REGION Network 11: Motor Conveyor Labeller
   RUNG wire#powerrail
      Contact( "Flag Motor" )
      Coil( "Motor" )
   END_RUNG
   // the same network as SCL:
   "Motor" := "Flag Motor";
END_REGION

REGION Network 12: Start Markem Input
   RUNG wire#powerrail
      Contact( "Flag Imaje Start" )
      Coil( "Imaje Output Start" )
   END_RUNG
   // the same network as SCL:
   "Imaje Output Start" := "Flag Imaje Start";
END_REGION

REGION Network 13: Pause Markem Input
   RUNG wire#powerrail
      Contact( "Flag Imaje Pause" )
      Coil( "Imaje Output Pause" )
   END_RUNG
   // the same network as SCL:
   "Imaje Output Pause" := "Flag Imaje Pause";
END_REGION

REGION Network 14: Trigger Markem Stamp
   RUNG wire#powerrail
      Contact( "Flag Imaje Trigger" )
      Coil( "Imaje Output Trigger" )
   END_RUNG
   // the same network as SCL:
   "Imaje Output Trigger" := "Flag Imaje Trigger";
END_REGION

REGION Network 15: Mesin Sebelumnya
   RUNG wire#powerrail
      Contact( "Machine Running" )
      Coil( "Trigger Mesin Sebelumnya" )
   END_RUNG
   // the same network as SCL:
   "Trigger Mesin Sebelumnya" := "Machine Running";
END_REGION

REGION Network 16: Error Output
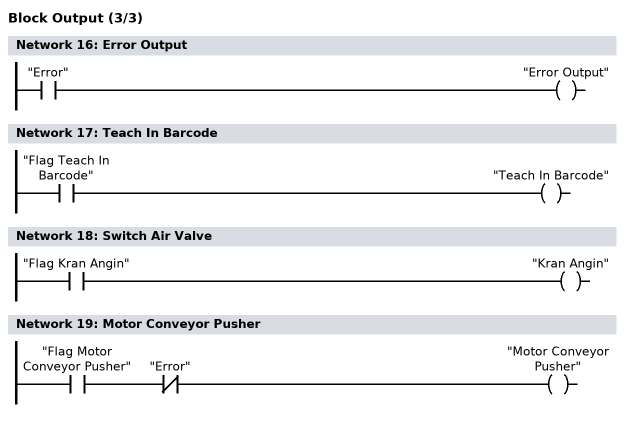
   RUNG wire#powerrail
      Contact( "Error" )
      Coil( "Error Output" )
   END_RUNG
   // the same network as SCL:
   "Error Output" := "Error";
END_REGION

REGION Network 17: Teach In Barcode
   RUNG wire#powerrail
      Contact( "Flag Teach In Barcode" )
      Coil( "Teach In Barcode" )
   END_RUNG
   // the same network as SCL:
   "Teach In Barcode" := "Flag Teach In Barcode";
END_REGION

REGION Network 18: Switch Air Valve
   RUNG wire#powerrail
      Contact( "Flag Kran Angin" )
      Coil( "Kran Angin" )
   END_RUNG
   // the same network as SCL:
   "Kran Angin" := "Flag Kran Angin";
END_REGION

REGION Network 19: Motor Conveyor Pusher
   RUNG wire#powerrail
      Contact( "Flag Motor Conveyor Pusher" )
      I_Contact( "Error" )
      Coil( "Motor Conveyor Pusher" )
   END_RUNG
   // the same network as SCL:
   "Motor Conveyor Pusher" := "Flag Motor Conveyor Pusher" AND NOT "Error";
END_REGION

REGION Network 20: Motor Heating Roll
END_REGION
END_FUNCTION_BLOCK

FUNCTION_BLOCK "S Block Current Shift"   // FB4, LAD
{ S7_Optimized_Access := 'TRUE' }
VERSION : 0.1
   VAR_TEMP   // added for the SCL form of the ladder/FBD networks
      _w1 : Bool;
      _w2 : Bool;
   END_VAR
BEGIN

REGION Network 1: Input Sloft ........................................................................page 1
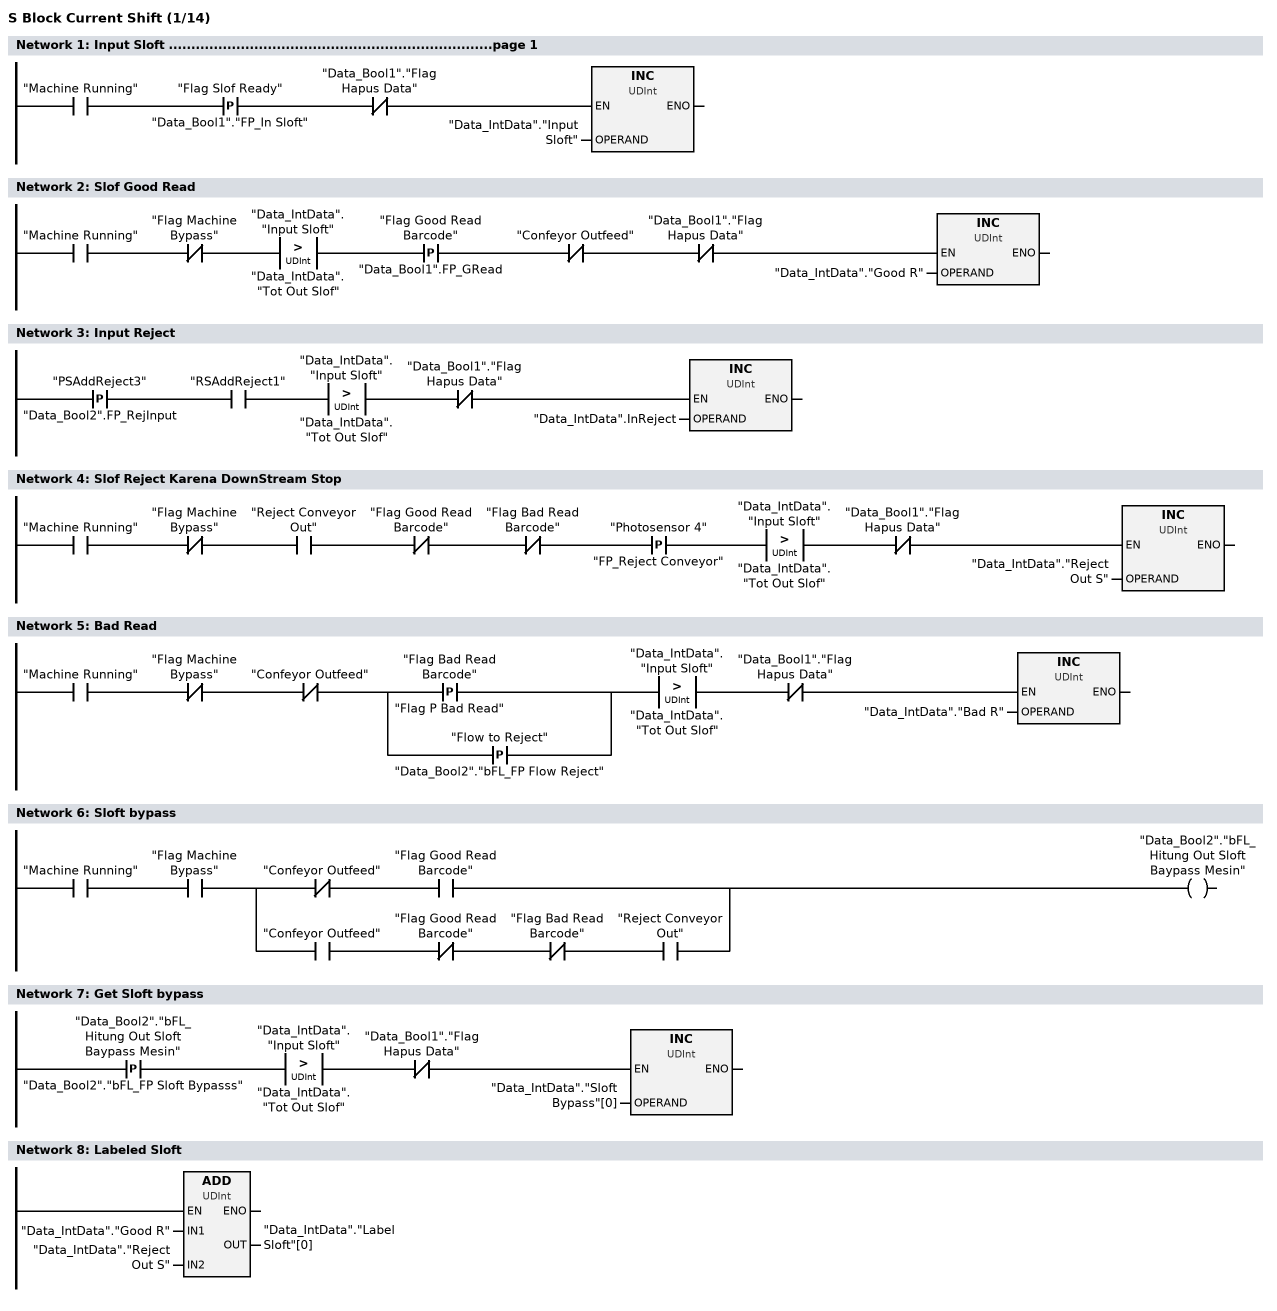
   RUNG wire#powerrail
      Contact( "Machine Running" )
      P_Contact(operand := "Flag Slof Ready", bit := "Data_Bool1"."FP_In Sloft")
      I_Contact( "Data_Bool1"."Flag Hapus Data" )
      { S7_Templates := "DestType := UDInt"; S7_GenerateENO := "TRUE" } Inc( "Data_IntData"."Input Sloft" )
   END_RUNG
   // the same network as SCL:
   #_w1 := "Machine Running" AND "Flag Slof Ready" AND NOT "Data_Bool1"."FP_In Sloft";   // rising edge of "Flag Slof Ready"
   "Data_Bool1"."FP_In Sloft" := "Flag Slof Ready";
   IF #_w1 AND NOT "Data_Bool1"."Flag Hapus Data" THEN
       "Data_IntData"."Input Sloft" := "Data_IntData"."Input Sloft" + 1;
   END_IF;
END_REGION

REGION Network 2: Slof Good Read
   RUNG wire#powerrail
      Contact( "Machine Running" )
      I_Contact( "Flag Machine Bypass" )
      { S7_Templates := "SrcType := UDInt" } GT_Contact(in1 := "Data_IntData"."Input Sloft", in2 := "Data_IntData"."Tot Out Slof")
      P_Contact(operand := "Flag Good Read Barcode", bit := "Data_Bool1".FP_GRead)
      I_Contact( "Confeyor Outfeed" )
      I_Contact( "Data_Bool1"."Flag Hapus Data" )
      { S7_Templates := "DestType := UDInt"; S7_GenerateENO := "TRUE" } Inc( "Data_IntData"."Good R" )
   END_RUNG
   // the same network as SCL:
   #_w1 := "Machine Running" AND NOT "Flag Machine Bypass" AND ("Data_IntData"."Input Sloft" > "Data_IntData"."Tot Out Slof") AND "Flag Good Read Barcode" AND NOT "Data_Bool1".FP_GRead;   // rising edge of "Flag Good Read Barcode"
   "Data_Bool1".FP_GRead := "Flag Good Read Barcode";
   IF #_w1 AND NOT "Confeyor Outfeed" AND NOT "Data_Bool1"."Flag Hapus Data" THEN
       "Data_IntData"."Good R" := "Data_IntData"."Good R" + 1;
   END_IF;
END_REGION

REGION Network 3: Input Reject
   RUNG wire#powerrail
      P_Contact(operand := "PSAddReject3", bit := "Data_Bool2".FP_RejInput)
      Contact( "RSAddReject1" )
      { S7_Templates := "SrcType := UDInt" } GT_Contact(in1 := "Data_IntData"."Input Sloft", in2 := "Data_IntData"."Tot Out Slof")
      I_Contact( "Data_Bool1"."Flag Hapus Data" )
      { S7_Templates := "DestType := UDInt"; S7_GenerateENO := "TRUE" } Inc( "Data_IntData".InReject )
   END_RUNG
   // the same network as SCL:
   #_w1 := "PSAddReject3" AND NOT "Data_Bool2".FP_RejInput;   // rising edge of "PSAddReject3"
   "Data_Bool2".FP_RejInput := "PSAddReject3";
   IF #_w1 AND "RSAddReject1" AND ("Data_IntData"."Input Sloft" > "Data_IntData"."Tot Out Slof") AND NOT "Data_Bool1"."Flag Hapus Data" THEN
       "Data_IntData".InReject := "Data_IntData".InReject + 1;
   END_IF;
END_REGION

REGION Network 4: Slof Reject Karena DownStream Stop
   RUNG wire#powerrail
      Contact( "Machine Running" )
      I_Contact( "Flag Machine Bypass" )
      Contact( "Reject Conveyor Out" )
      I_Contact( "Flag Good Read Barcode" )
      I_Contact( "Flag Bad Read Barcode" )
      P_Contact(operand := "Photosensor 4", bit := "FP_Reject Conveyor")
      { S7_Templates := "SrcType := UDInt" } GT_Contact(in1 := "Data_IntData"."Input Sloft", in2 := "Data_IntData"."Tot Out Slof")
      I_Contact( "Data_Bool1"."Flag Hapus Data" )
      { S7_Templates := "DestType := UDInt"; S7_GenerateENO := "TRUE" } Inc( "Data_IntData"."Reject Out S" )
   END_RUNG
   // the same network as SCL:
   #_w1 := "Machine Running" AND NOT "Flag Machine Bypass" AND "Reject Conveyor Out" AND NOT "Flag Good Read Barcode" AND NOT "Flag Bad Read Barcode" AND "Photosensor 4" AND NOT "FP_Reject Conveyor";   // rising edge of "Photosensor 4"
   "FP_Reject Conveyor" := "Photosensor 4";
   IF #_w1 AND ("Data_IntData"."Input Sloft" > "Data_IntData"."Tot Out Slof") AND NOT "Data_Bool1"."Flag Hapus Data" THEN
       "Data_IntData"."Reject Out S" := "Data_IntData"."Reject Out S" + 1;
   END_IF;
END_REGION

REGION Network 5: Bad Read
   RUNG wire#powerrail
      Contact( "Machine Running" )
      I_Contact( "Flag Machine Bypass" )
      I_Contact( "Confeyor Outfeed" )
      wire#w1
      P_Contact(operand := "Flag Bad Read Barcode", bit := "Flag P Bad Read")
      wire#w2
      { S7_Templates := "SrcType := UDInt" } GT_Contact(in1 := "Data_IntData"."Input Sloft", in2 := "Data_IntData"."Tot Out Slof")
      I_Contact( "Data_Bool1"."Flag Hapus Data" )
      { S7_Templates := "DestType := UDInt"; S7_GenerateENO := "TRUE" } Inc( "Data_IntData"."Bad R" )
   END_RUNG
   RUNG wire#w1
      P_Contact(operand := "Flow to Reject", bit := "Data_Bool2"."bFL_FP Flow Reject")
   END_RUNG wire#w2
   // the same network as SCL:
   #_w1 := "Machine Running" AND NOT "Flag Machine Bypass" AND NOT "Confeyor Outfeed" AND "Flag Bad Read Barcode" AND NOT "Flag P Bad Read";   // rising edge of "Flag Bad Read Barcode"
   "Flag P Bad Read" := "Flag Bad Read Barcode";
   #_w2 := "Machine Running" AND NOT "Flag Machine Bypass" AND NOT "Confeyor Outfeed" AND "Flow to Reject" AND NOT "Data_Bool2"."bFL_FP Flow Reject";   // rising edge of "Flow to Reject"
   "Data_Bool2"."bFL_FP Flow Reject" := "Flow to Reject";
   IF (#_w1 OR #_w2) AND ("Data_IntData"."Input Sloft" > "Data_IntData"."Tot Out Slof") AND NOT "Data_Bool1"."Flag Hapus Data" THEN
       "Data_IntData"."Bad R" := "Data_IntData"."Bad R" + 1;
   END_IF;
END_REGION

REGION Network 6: Sloft bypass
   RUNG wire#powerrail
      Contact( "Machine Running" )
      Contact( "Flag Machine Bypass" )
      wire#w1
      I_Contact( "Confeyor Outfeed" )
      Contact( "Flag Good Read Barcode" )
      wire#w2
      Coil( "Data_Bool2"."bFL_Hitung Out Sloft Baypass Mesin" )
   END_RUNG
   RUNG wire#w1
      Contact( "Confeyor Outfeed" )
      I_Contact( "Flag Good Read Barcode" )
      I_Contact( "Flag Bad Read Barcode" )
      Contact( "Reject Conveyor Out" )
   END_RUNG wire#w2
   // the same network as SCL:
   "Data_Bool2"."bFL_Hitung Out Sloft Baypass Mesin" := "Machine Running" AND "Flag Machine Bypass" AND ((NOT "Confeyor Outfeed" AND "Flag Good Read Barcode") OR ("Confeyor Outfeed" AND NOT "Flag Good Read Barcode" AND NOT "Flag Bad Read Barcode" AND "Reject Conveyor Out"));
END_REGION

REGION Network 7: Get Sloft bypass
   RUNG wire#powerrail
      P_Contact(operand := "Data_Bool2"."bFL_Hitung Out Sloft Baypass Mesin", bit := "Data_Bool2"."bFL_FP Sloft Bypasss")
      { S7_Templates := "SrcType := UDInt" } GT_Contact(in1 := "Data_IntData"."Input Sloft", in2 := "Data_IntData"."Tot Out Slof")
      I_Contact( "Data_Bool1"."Flag Hapus Data" )
      { S7_Templates := "DestType := UDInt"; S7_GenerateENO := "TRUE" } Inc( "Data_IntData"."Sloft Bypass"[0] )
   END_RUNG
   // the same network as SCL:
   #_w1 := "Data_Bool2"."bFL_Hitung Out Sloft Baypass Mesin" AND NOT "Data_Bool2"."bFL_FP Sloft Bypasss";   // rising edge of "Data_Bool2"."bFL_Hitung Out Sloft Baypass Mesin"
   "Data_Bool2"."bFL_FP Sloft Bypasss" := "Data_Bool2"."bFL_Hitung Out Sloft Baypass Mesin";
   IF #_w1 AND ("Data_IntData"."Input Sloft" > "Data_IntData"."Tot Out Slof") AND NOT "Data_Bool1"."Flag Hapus Data" THEN
       "Data_IntData"."Sloft Bypass"[0] := "Data_IntData"."Sloft Bypass"[0] + 1;
   END_IF;
END_REGION

REGION Network 8: Labeled Sloft
   RUNG wire#powerrail
      { S7_Templates := "SrcType := UDInt"; S7_GenerateENO := "TRUE" } Add(in1 := "Data_IntData"."Good R", in2 := "Data_IntData"."Reject Out S", out => "Data_IntData"."Label Sloft"[0])
   END_RUNG
   // the same network as SCL:
   "Data_IntData"."Label Sloft"[0] := "Data_IntData"."Good R" + "Data_IntData"."Reject Out S";
END_REGION

REGION Network 9: Unlabeled Sloft
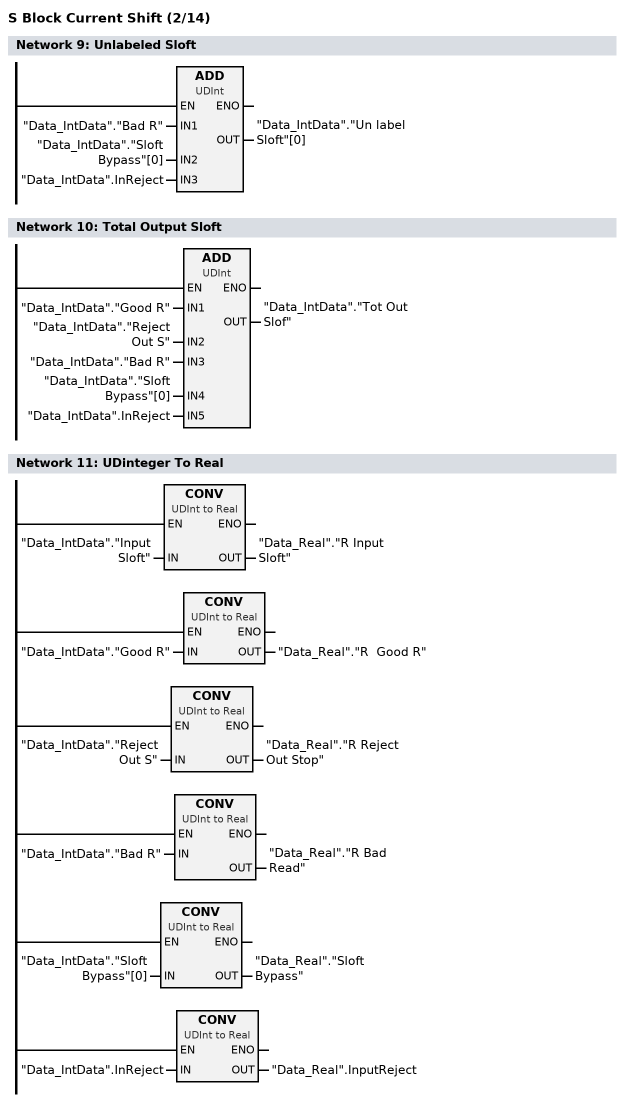
   RUNG wire#powerrail
      { S7_Templates := "SrcType := UDInt"; S7_GenerateENO := "TRUE" } Add(in1 := "Data_IntData"."Bad R", in2 := "Data_IntData"."Sloft Bypass"[0], in3 := "Data_IntData".InReject, out => "Data_IntData"."Un label Sloft"[0])
   END_RUNG
   // the same network as SCL:
   "Data_IntData"."Un label Sloft"[0] := "Data_IntData"."Bad R" + "Data_IntData"."Sloft Bypass"[0] + "Data_IntData".InReject;
END_REGION

REGION Network 10: Total Output Sloft
   RUNG wire#powerrail
      { S7_Templates := "SrcType := UDInt"; S7_GenerateENO := "TRUE" } Add(in1 := "Data_IntData"."Good R", in2 := "Data_IntData"."Reject Out S", in3 := "Data_IntData"."Bad R", in4 := "Data_IntData"."Sloft Bypass"[0], in5 := "Data_IntData".InReject, out => "Data_IntData"."Tot Out Slof")
   END_RUNG
   // the same network as SCL:
   "Data_IntData"."Tot Out Slof" := "Data_IntData"."Good R" + "Data_IntData"."Reject Out S" + "Data_IntData"."Bad R" + "Data_IntData"."Sloft Bypass"[0] + "Data_IntData".InReject;
END_REGION

REGION Network 11: UDinteger To Real
   RUNG wire#powerrail
      { S7_Templates := "[SrcType := UDInt, DestType := Real]"; S7_GenerateENO := "TRUE" } Convert(in := "Data_IntData"."Input Sloft", out => "Data_Real"."R Input Sloft")
   END_RUNG
   RUNG wire#powerrail
      { S7_Templates := "[SrcType := UDInt, DestType := Real]"; S7_GenerateENO := "TRUE" } Convert(in := "Data_IntData"."Good R", out => "Data_Real"."R  Good R")
   END_RUNG
   RUNG wire#powerrail
      { S7_Templates := "[SrcType := UDInt, DestType := Real]"; S7_GenerateENO := "TRUE" } Convert(in := "Data_IntData"."Reject Out S", out => "Data_Real"."R Reject Out Stop")
   END_RUNG
   RUNG wire#powerrail
      { S7_Templates := "[SrcType := UDInt, DestType := Real]"; S7_GenerateENO := "TRUE" } Convert(in := "Data_IntData"."Bad R", out => "Data_Real"."R Bad Read")
   END_RUNG
   RUNG wire#powerrail
      { S7_Templates := "[SrcType := UDInt, DestType := Real]"; S7_GenerateENO := "TRUE" } Convert(in := "Data_IntData"."Sloft Bypass"[0], out => "Data_Real"."Sloft Bypass")
   END_RUNG
   RUNG wire#powerrail
      { S7_Templates := "[SrcType := UDInt, DestType := Real]"; S7_GenerateENO := "TRUE" } Convert(in := "Data_IntData".InReject, out => "Data_Real".InputReject)
   END_RUNG
   // the same network as SCL:
   "Data_Real"."R Input Sloft" := UDINT_TO_REAL("Data_IntData"."Input Sloft");
   "Data_Real"."R  Good R" := UDINT_TO_REAL("Data_IntData"."Good R");
   "Data_Real"."R Reject Out Stop" := UDINT_TO_REAL("Data_IntData"."Reject Out S");
   "Data_Real"."R Bad Read" := UDINT_TO_REAL("Data_IntData"."Bad R");
   "Data_Real"."Sloft Bypass" := UDINT_TO_REAL("Data_IntData"."Sloft Bypass"[0]);
   "Data_Real".InputReject := UDINT_TO_REAL("Data_IntData".InReject);
END_REGION

REGION Network 12: % Sloft terhadap Input Sloft
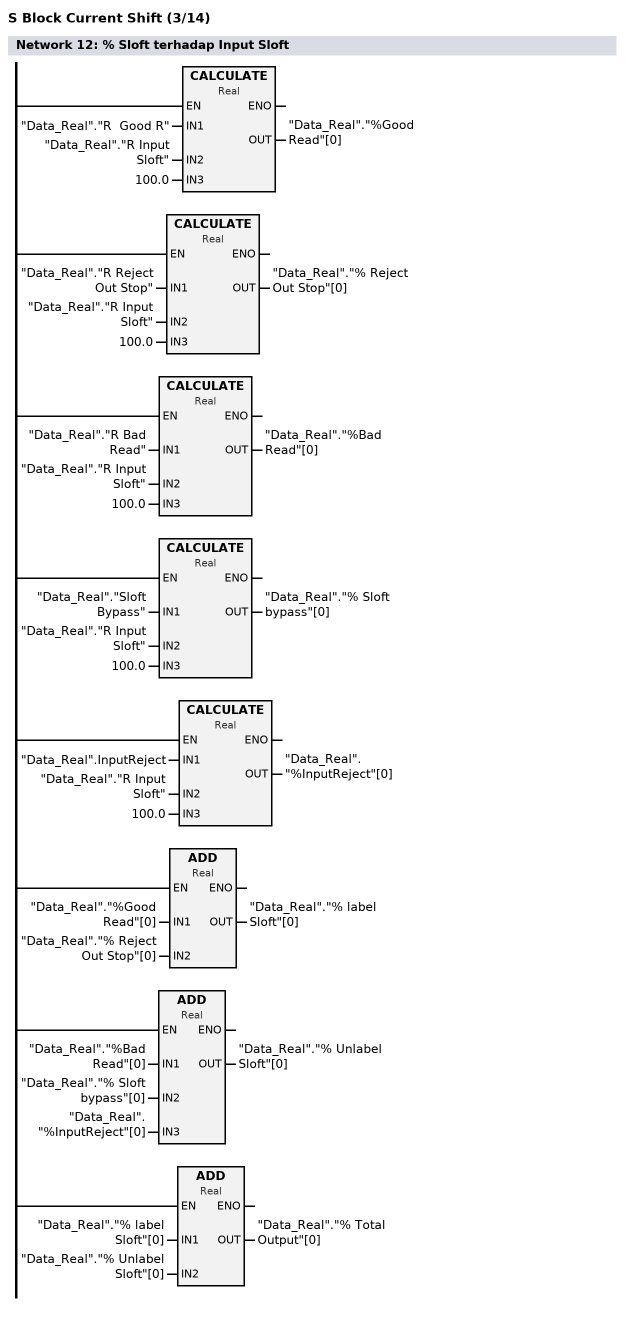
   RUNG wire#powerrail
      { S7_Templates := "SrcType := Real"; S7_GenerateENO := "TRUE"; S7_Expression := "(IN1/IN2)*IN3" } Calculate(in1 := "Data_Real"."R  Good R", in2 := "Data_Real"."R Input Sloft", in3 := 100.0, out => "Data_Real"."%Good Read"[0])
   END_RUNG
   RUNG wire#powerrail
      { S7_Templates := "SrcType := Real"; S7_GenerateENO := "TRUE"; S7_Expression := "(IN1/IN2)*IN3" } Calculate(in1 := "Data_Real"."R Reject Out Stop", in2 := "Data_Real"."R Input Sloft", in3 := 100.0, out => "Data_Real"."% Reject Out Stop"[0])
   END_RUNG
   RUNG wire#powerrail
      { S7_Templates := "SrcType := Real"; S7_GenerateENO := "TRUE"; S7_Expression := "(IN1/IN2)*IN3" } Calculate(in1 := "Data_Real"."R Bad Read", in2 := "Data_Real"."R Input Sloft", in3 := 100.0, out => "Data_Real"."%Bad Read"[0])
   END_RUNG
   RUNG wire#powerrail
      { S7_Templates := "SrcType := Real"; S7_GenerateENO := "TRUE"; S7_Expression := "(IN1/IN2)*IN3" } Calculate(in1 := "Data_Real"."Sloft Bypass", in2 := "Data_Real"."R Input Sloft", in3 := 100.0, out => "Data_Real"."% Sloft bypass"[0])
   END_RUNG
   RUNG wire#powerrail
      { S7_Templates := "SrcType := Real"; S7_GenerateENO := "TRUE"; S7_Expression := "(IN1/IN2)*IN3" } Calculate(in1 := "Data_Real".InputReject, in2 := "Data_Real"."R Input Sloft", in3 := 100.0, out => "Data_Real"."%InputReject"[0])
   END_RUNG
   RUNG wire#powerrail
      { S7_Templates := "SrcType := Real"; S7_GenerateENO := "TRUE" } Add(in1 := "Data_Real"."%Good Read"[0], in2 := "Data_Real"."% Reject Out Stop"[0], out => "Data_Real"."% label Sloft"[0])
   END_RUNG
   RUNG wire#powerrail
      { S7_Templates := "SrcType := Real"; S7_GenerateENO := "TRUE" } Add(in1 := "Data_Real"."%Bad Read"[0], in2 := "Data_Real"."% Sloft bypass"[0], in3 := "Data_Real"."%InputReject"[0], out => "Data_Real"."% Unlabel Sloft"[0])
   END_RUNG
   RUNG wire#powerrail
      { S7_Templates := "SrcType := Real"; S7_GenerateENO := "TRUE" } Add(in1 := "Data_Real"."% label Sloft"[0], in2 := "Data_Real"."% Unlabel Sloft"[0], out => "Data_Real"."% Total Output"[0])
   END_RUNG
   // the same network as SCL:
   "Data_Real"."%Good Read"[0] := ("Data_Real"."R  Good R"/"Data_Real"."R Input Sloft")*100.0;
   "Data_Real"."% Reject Out Stop"[0] := ("Data_Real"."R Reject Out Stop"/"Data_Real"."R Input Sloft")*100.0;
   "Data_Real"."%Bad Read"[0] := ("Data_Real"."R Bad Read"/"Data_Real"."R Input Sloft")*100.0;
   "Data_Real"."% Sloft bypass"[0] := ("Data_Real"."Sloft Bypass"/"Data_Real"."R Input Sloft")*100.0;
   "Data_Real"."%InputReject"[0] := ("Data_Real".InputReject/"Data_Real"."R Input Sloft")*100.0;
   "Data_Real"."% label Sloft"[0] := "Data_Real"."%Good Read"[0] + "Data_Real"."% Reject Out Stop"[0];
   "Data_Real"."% Unlabel Sloft"[0] := "Data_Real"."%Bad Read"[0] + "Data_Real"."% Sloft bypass"[0] + "Data_Real"."%InputReject"[0];
   "Data_Real"."% Total Output"[0] := "Data_Real"."% label Sloft"[0] + "Data_Real"."% Unlabel Sloft"[0];
END_REGION

REGION Network 13: ----------- Get Image Output Trigger
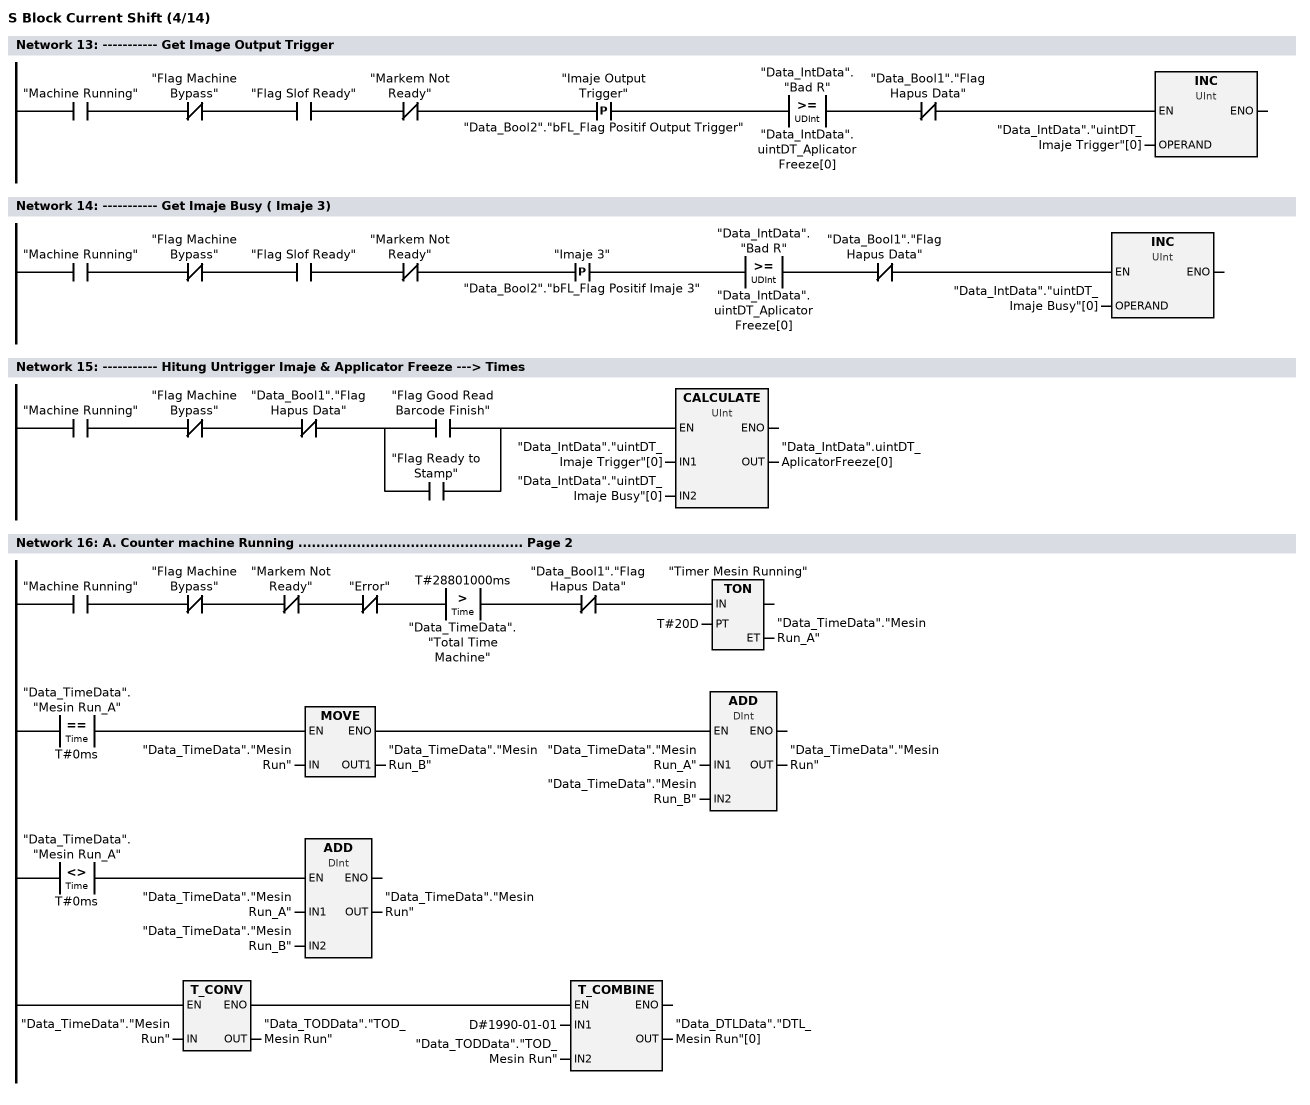
   RUNG wire#powerrail
      Contact( "Machine Running" )
      I_Contact( "Flag Machine Bypass" )
      Contact( "Flag Slof Ready" )
      I_Contact( "Markem Not Ready" )
      P_Contact(operand := "Imaje Output Trigger", bit := "Data_Bool2"."bFL_Flag Positif Output Trigger")
      { S7_Templates := "SrcType := UDInt" } GE_Contact(in1 := "Data_IntData"."Bad R", in2 := "Data_IntData".uintDT_AplicatorFreeze[0])
      I_Contact( "Data_Bool1"."Flag Hapus Data" )
      { S7_Templates := "DestType := UInt"; S7_GenerateENO := "TRUE" } Inc( "Data_IntData"."uintDT_Imaje Trigger"[0] )
   END_RUNG
   // the same network as SCL:
   #_w1 := "Machine Running" AND NOT "Flag Machine Bypass" AND "Flag Slof Ready" AND NOT "Markem Not Ready" AND "Imaje Output Trigger" AND NOT "Data_Bool2"."bFL_Flag Positif Output Trigger";   // rising edge of "Imaje Output Trigger"
   "Data_Bool2"."bFL_Flag Positif Output Trigger" := "Imaje Output Trigger";
   IF #_w1 AND ("Data_IntData"."Bad R" >= "Data_IntData".uintDT_AplicatorFreeze[0]) AND NOT "Data_Bool1"."Flag Hapus Data" THEN
       "Data_IntData"."uintDT_Imaje Trigger"[0] := "Data_IntData"."uintDT_Imaje Trigger"[0] + 1;
   END_IF;
END_REGION

REGION Network 14: ----------- Get Imaje Busy ( Imaje 3)
   RUNG wire#powerrail
      Contact( "Machine Running" )
      I_Contact( "Flag Machine Bypass" )
      Contact( "Flag Slof Ready" )
      I_Contact( "Markem Not Ready" )
      P_Contact(operand := "Imaje 3", bit := "Data_Bool2"."bFL_Flag Positif Imaje 3")
      { S7_Templates := "SrcType := UDInt" } GE_Contact(in1 := "Data_IntData"."Bad R", in2 := "Data_IntData".uintDT_AplicatorFreeze[0])
      I_Contact( "Data_Bool1"."Flag Hapus Data" )
      { S7_Templates := "DestType := UInt"; S7_GenerateENO := "TRUE" } Inc( "Data_IntData"."uintDT_Imaje Busy"[0] )
   END_RUNG
   // the same network as SCL:
   #_w1 := "Machine Running" AND NOT "Flag Machine Bypass" AND "Flag Slof Ready" AND NOT "Markem Not Ready" AND "Imaje 3" AND NOT "Data_Bool2"."bFL_Flag Positif Imaje 3";   // rising edge of "Imaje 3"
   "Data_Bool2"."bFL_Flag Positif Imaje 3" := "Imaje 3";
   IF #_w1 AND ("Data_IntData"."Bad R" >= "Data_IntData".uintDT_AplicatorFreeze[0]) AND NOT "Data_Bool1"."Flag Hapus Data" THEN
       "Data_IntData"."uintDT_Imaje Busy"[0] := "Data_IntData"."uintDT_Imaje Busy"[0] + 1;
   END_IF;
END_REGION

REGION Network 15: ----------- Hitung Untrigger Imaje & Applicator Freeze ---> Times
   RUNG wire#powerrail
      Contact( "Machine Running" )
      I_Contact( "Flag Machine Bypass" )
      I_Contact( "Data_Bool1"."Flag Hapus Data" )
      wire#w1
      Contact( "Flag Good Read Barcode Finish" )
      wire#w2
      { S7_Templates := "SrcType := UInt"; S7_GenerateENO := "TRUE"; S7_Expression := "IN1- IN2" } Calculate(in1 := "Data_IntData"."uintDT_Imaje Trigger"[0], in2 := "Data_IntData"."uintDT_Imaje Busy"[0], out => "Data_IntData".uintDT_AplicatorFreeze[0])
   END_RUNG
   RUNG wire#w1
      Contact( "Flag Ready to Stamp" )
   END_RUNG wire#w2
   // the same network as SCL:
   IF "Machine Running" AND NOT "Flag Machine Bypass" AND NOT "Data_Bool1"."Flag Hapus Data" AND ("Flag Good Read Barcode Finish" OR "Flag Ready to Stamp") THEN
       "Data_IntData".uintDT_AplicatorFreeze[0] := "Data_IntData"."uintDT_Imaje Trigger"[0]- "Data_IntData"."uintDT_Imaje Busy"[0];
   END_IF;
END_REGION

REGION Network 16: A. Counter machine Running .................................................. Page 2
   // ENO of a box is taken as its EN; it also drops when the box reports an error
   "Timer Mesin Running".TON(IN := "Machine Running" AND NOT "Flag Machine Bypass" AND NOT "Markem Not Ready" AND NOT "Error" AND (T#28801000ms > "Data_TimeData"."Total Time Machine") AND NOT "Data_Bool1"."Flag Hapus Data",
                           PT := T#20D,
                           ET => "Data_TimeData"."Mesin Run_A");
   IF "Data_TimeData"."Mesin Run_A" = T#0ms THEN
       "Data_TimeData"."Mesin Run_B" := "Data_TimeData"."Mesin Run";
       "Data_TimeData"."Mesin Run" := "Data_TimeData"."Mesin Run_A" + "Data_TimeData"."Mesin Run_B";
   END_IF;
   IF "Data_TimeData"."Mesin Run_A" <> T#0ms THEN
       "Data_TimeData"."Mesin Run" := "Data_TimeData"."Mesin Run_A" + "Data_TimeData"."Mesin Run_B";
   END_IF;
   "Data_TODData"."TOD_Mesin Run" := T_CONV(IN := "Data_TimeData"."Mesin Run");
   "Data_DTLData"."DTL_Mesin Run"[0] := T_COMBINE(IN1 := D#1990-01-01, IN2 := "Data_TODData"."TOD_Mesin Run");
END_REGION

REGION Network 17: B. Counter machine Running Baypass Stamp
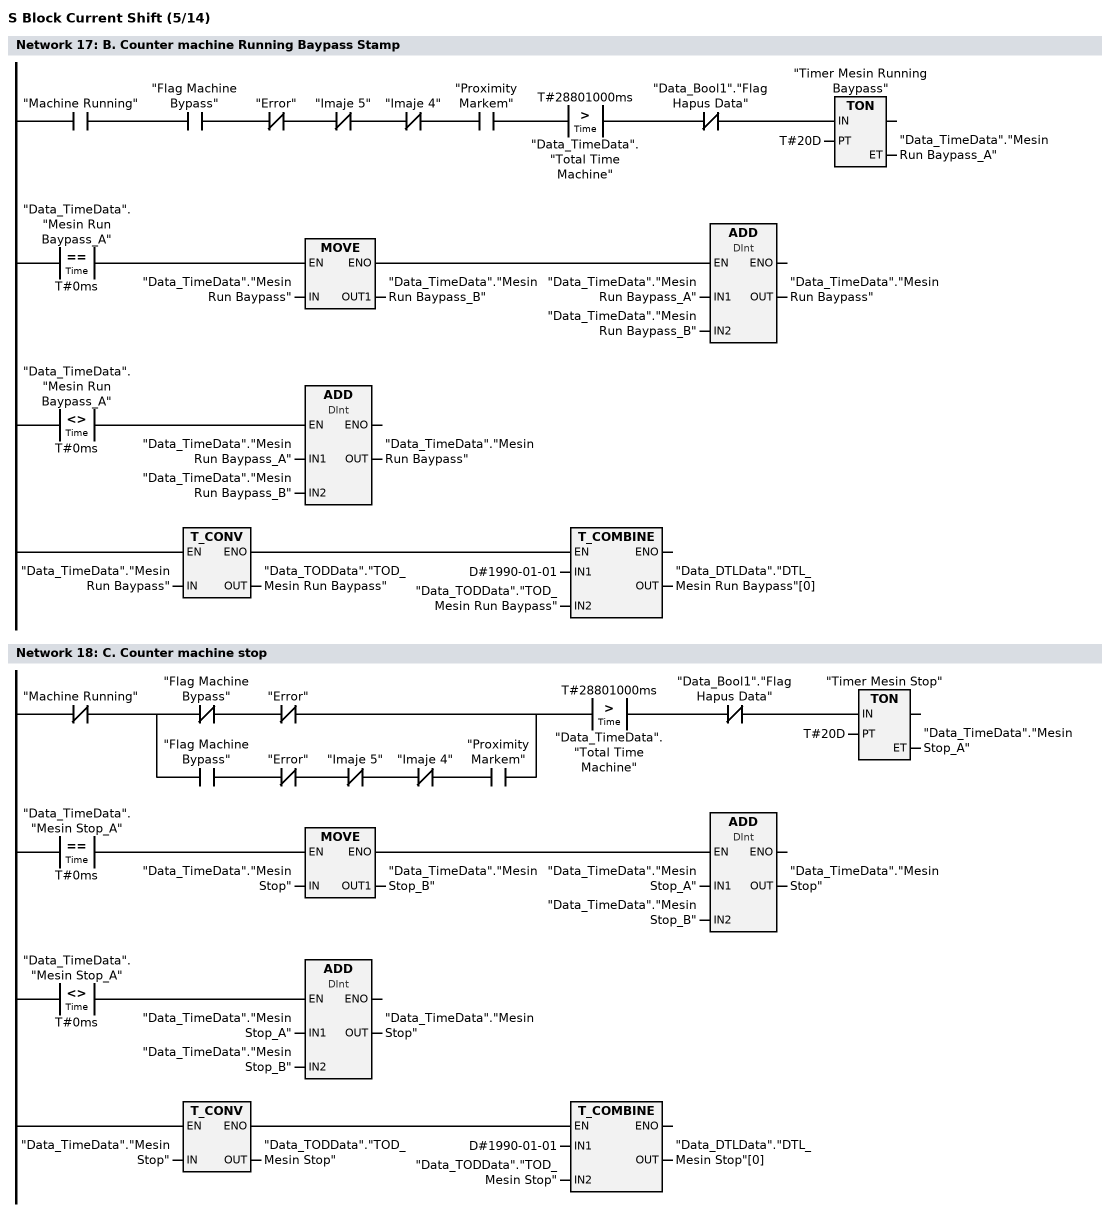
   // ENO of a box is taken as its EN; it also drops when the box reports an error
   "Timer Mesin Running Baypass".TON(IN := "Machine Running" AND "Flag Machine Bypass" AND NOT "Error" AND NOT "Imaje 5" AND NOT "Imaje 4" AND "Proximity Markem" AND (T#28801000ms > "Data_TimeData"."Total Time Machine") AND NOT "Data_Bool1"."Flag Hapus Data",
                           PT := T#20D,
                           ET => "Data_TimeData"."Mesin Run Baypass_A");
   IF "Data_TimeData"."Mesin Run Baypass_A" = T#0ms THEN
       "Data_TimeData"."Mesin Run Baypass_B" := "Data_TimeData"."Mesin Run Baypass";
       "Data_TimeData"."Mesin Run Baypass" := "Data_TimeData"."Mesin Run Baypass_A" + "Data_TimeData"."Mesin Run Baypass_B";
   END_IF;
   IF "Data_TimeData"."Mesin Run Baypass_A" <> T#0ms THEN
       "Data_TimeData"."Mesin Run Baypass" := "Data_TimeData"."Mesin Run Baypass_A" + "Data_TimeData"."Mesin Run Baypass_B";
   END_IF;
   "Data_TODData"."TOD_Mesin Run Baypass" := T_CONV(IN := "Data_TimeData"."Mesin Run Baypass");
   "Data_DTLData"."DTL_Mesin Run Baypass"[0] := T_COMBINE(IN1 := D#1990-01-01,
                           IN2 := "Data_TODData"."TOD_Mesin Run Baypass");
END_REGION

REGION Network 18: C. Counter machine stop
   // ENO of a box is taken as its EN; it also drops when the box reports an error
   "Timer Mesin Stop".TON(IN := NOT "Machine Running" AND ((NOT "Flag Machine Bypass" AND NOT "Error") OR ("Flag Machine Bypass" AND NOT "Error" AND NOT "Imaje 5" AND NOT "Imaje 4" AND "Proximity Markem")) AND (T#28801000ms > "Data_TimeData"."Total Time Machine") AND NOT "Data_Bool1"."Flag Hapus Data",
                          PT := T#20D,
                          ET => "Data_TimeData"."Mesin Stop_A");
   IF "Data_TimeData"."Mesin Stop_A" = T#0ms THEN
       "Data_TimeData"."Mesin Stop_B" := "Data_TimeData"."Mesin Stop";
       "Data_TimeData"."Mesin Stop" := "Data_TimeData"."Mesin Stop_A" + "Data_TimeData"."Mesin Stop_B";
   END_IF;
   IF "Data_TimeData"."Mesin Stop_A" <> T#0ms THEN
       "Data_TimeData"."Mesin Stop" := "Data_TimeData"."Mesin Stop_A" + "Data_TimeData"."Mesin Stop_B";
   END_IF;
   "Data_TODData"."TOD_Mesin Stop" := T_CONV(IN := "Data_TimeData"."Mesin Stop");
   "Data_DTLData"."DTL_Mesin Stop"[0] := T_COMBINE(IN1 := D#1990-01-01, IN2 := "Data_TODData"."TOD_Mesin Stop");
END_REGION

REGION Network 19: D. Counter Machine Error
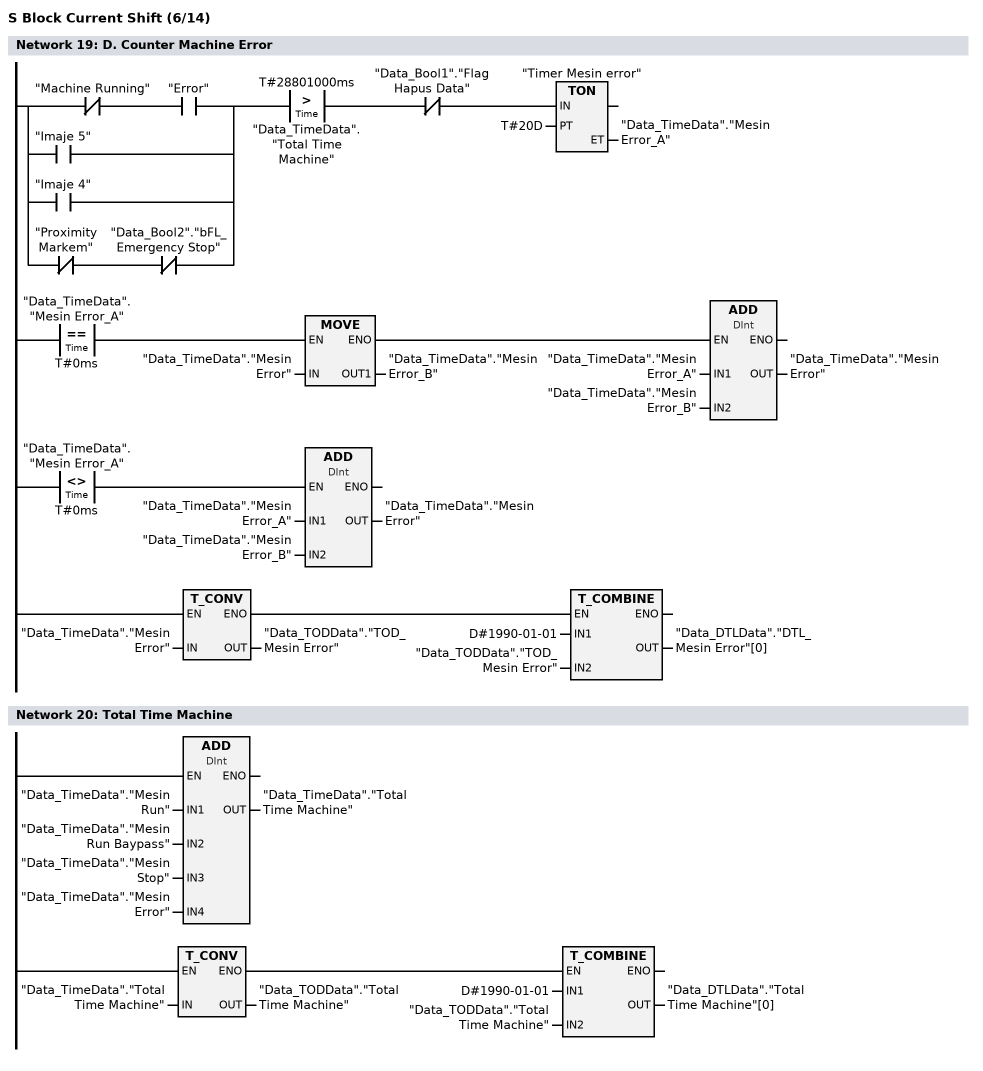
   // ENO of a box is taken as its EN; it also drops when the box reports an error
   "Timer Mesin error".TON(IN := ((NOT "Machine Running" AND "Error") OR "Imaje 5" OR "Imaje 4" OR (NOT "Proximity Markem" AND NOT "Data_Bool2"."bFL_Emergency Stop")) AND (T#28801000ms > "Data_TimeData"."Total Time Machine") AND NOT "Data_Bool1"."Flag Hapus Data",
                           PT := T#20D,
                           ET => "Data_TimeData"."Mesin Error_A");
   IF "Data_TimeData"."Mesin Error_A" = T#0ms THEN
       "Data_TimeData"."Mesin Error_B" := "Data_TimeData"."Mesin Error";
       "Data_TimeData"."Mesin Error" := "Data_TimeData"."Mesin Error_A" + "Data_TimeData"."Mesin Error_B";
   END_IF;
   IF "Data_TimeData"."Mesin Error_A" <> T#0ms THEN
       "Data_TimeData"."Mesin Error" := "Data_TimeData"."Mesin Error_A" + "Data_TimeData"."Mesin Error_B";
   END_IF;
   "Data_TODData"."TOD_Mesin Error" := T_CONV(IN := "Data_TimeData"."Mesin Error");
   "Data_DTLData"."DTL_Mesin Error"[0] := T_COMBINE(IN1 := D#1990-01-01,
                           IN2 := "Data_TODData"."TOD_Mesin Error");
END_REGION
